REGION Network 141
   RUNG wire#powerrail
      Contact( "Carrier_06_Status.9" )
      Coil( "EMS".Carrier[06].SDC_IN.EncoderCommFault )
   END_RUNG
   // the same network as SCL:
   "EMS".Carrier[06].SDC_IN.EncoderCommFault := "Carrier_06_Status.9";
END_REGION

REGION Network 142
   RUNG wire#powerrail
      Contact( "Carrier_06_Status.10" )
      Coil( "EMS".Carrier[06].SDC_IN.DriveCommFault )
   END_RUNG
   // the same network as SCL:
   "EMS".Carrier[06].SDC_IN.DriveCommFault := "Carrier_06_Status.10";
END_REGION

REGION Network 143
   RUNG wire#powerrail
      Contact( "Carrier_06_Status.11" )
      Coil( "EMS".Carrier[06].SDC_IN.HMICommFault )
   END_RUNG
   // the same network as SCL:
   "EMS".Carrier[06].SDC_IN.HMICommFault := "Carrier_06_Status.11";
END_REGION

REGION Network 144
   RUNG wire#powerrail
      Contact( "Carrier_06_Status.2" )
      Coil( "EMS".Carrier[06].SDC_IN.AutoMode )
   END_RUNG
   RUNG wire#powerrail
      Contact( "Carrier_06_Status.1" )
      Coil( "EMS".Carrier[06].SDC_IN.ManualMode )
   END_RUNG
   // the same network as SCL:
   "EMS".Carrier[06].SDC_IN.AutoMode := "Carrier_06_Status.2";
   "EMS".Carrier[06].SDC_IN.ManualMode := "Carrier_06_Status.1";
END_REGION

REGION Network 145
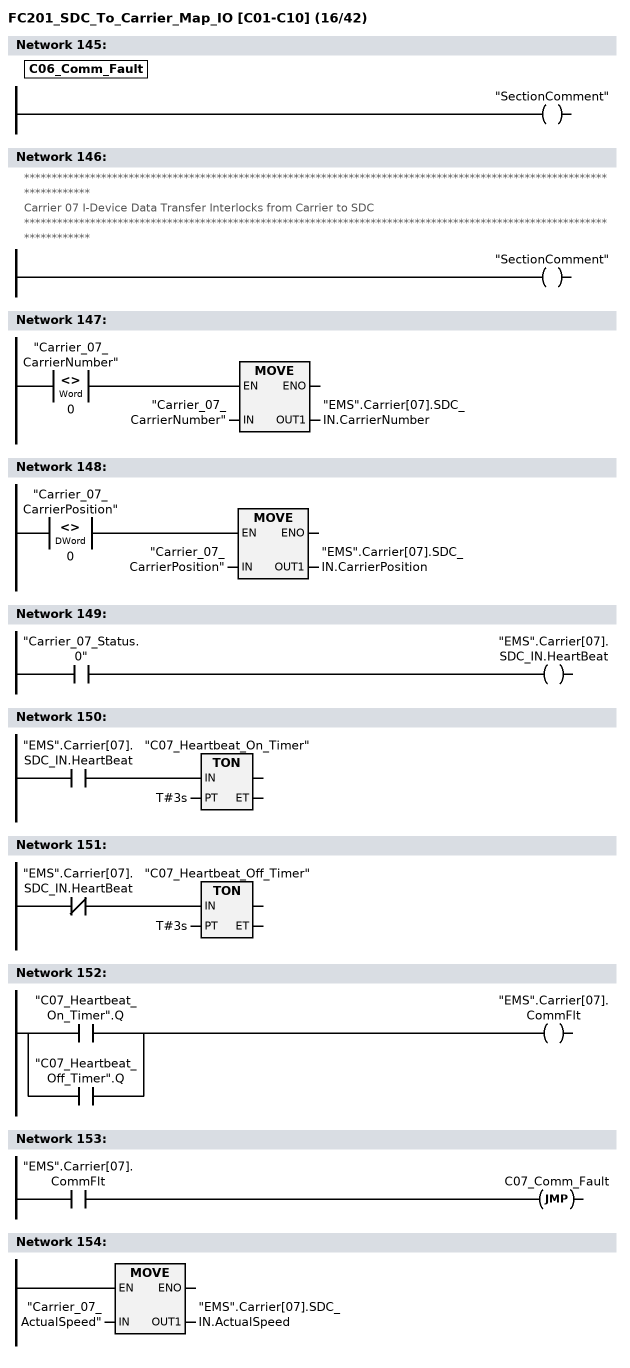
   Label( C06_Comm_Fault )
   RUNG wire#powerrail
      Coil( "SectionComment" )
   END_RUNG
   // the same network as SCL:
   C06_Comm_Fault:
   "SectionComment" := TRUE;
END_REGION

REGION Network 146
   // **********************************************************************************************************************
   // 
   // Carrier 07 I-Device Data Transfer Interlocks from Carrier to SDC
   // 
   // **********************************************************************************************************************
   RUNG wire#powerrail
      Coil( "SectionComment" )
   END_RUNG
   // the same network as SCL:
   "SectionComment" := TRUE;
END_REGION

REGION Network 147
   RUNG wire#powerrail
      { S7_Templates := "SrcType := Word" } NE_Contact(in1 := "Carrier_07_CarrierNumber", in2 := 0)
      Move(in := "Carrier_07_CarrierNumber", out1 => "EMS".Carrier[07].SDC_IN.CarrierNumber)
   END_RUNG
   // the same network as SCL:
   IF "Carrier_07_CarrierNumber" <> 0 THEN
       "EMS".Carrier[07].SDC_IN.CarrierNumber := "Carrier_07_CarrierNumber";
   END_IF;
END_REGION

REGION Network 148
   RUNG wire#powerrail
      { S7_Templates := "SrcType := DWord" } NE_Contact(in1 := "Carrier_07_CarrierPosition", in2 := 0)
      Move(in := "Carrier_07_CarrierPosition", out1 => "EMS".Carrier[07].SDC_IN.CarrierPosition)
   END_RUNG
   // the same network as SCL:
   IF "Carrier_07_CarrierPosition" <> 0 THEN
       "EMS".Carrier[07].SDC_IN.CarrierPosition := "Carrier_07_CarrierPosition";
   END_IF;
END_REGION

REGION Network 149
   RUNG wire#powerrail
      Contact( "Carrier_07_Status.0" )
      Coil( "EMS".Carrier[07].SDC_IN.HeartBeat )
   END_RUNG
   // the same network as SCL:
   "EMS".Carrier[07].SDC_IN.HeartBeat := "Carrier_07_Status.0";
END_REGION

REGION Network 150
   "C07_Heartbeat_On_Timer".TON(IN := "EMS".Carrier[07].SDC_IN.HeartBeat, PT := T#3s);
END_REGION

REGION Network 151
   "C07_Heartbeat_Off_Timer".TON(IN := NOT "EMS".Carrier[07].SDC_IN.HeartBeat, PT := T#3s);
END_REGION

REGION Network 152
   RUNG wire#powerrail
      Contact( "C07_Heartbeat_On_Timer".Q )
      wire#w1
      Coil( "EMS".Carrier[07].CommFlt )
   END_RUNG
   RUNG wire#powerrail
      Contact( "C07_Heartbeat_Off_Timer".Q )
   END_RUNG wire#w1
   // the same network as SCL:
   "EMS".Carrier[07].CommFlt := "C07_Heartbeat_On_Timer".Q OR "C07_Heartbeat_Off_Timer".Q;
END_REGION

REGION Network 153
   RUNG wire#powerrail
      Contact( "EMS".Carrier[07].CommFlt )
      JumpCoil( C07_Comm_Fault )
   END_RUNG
   // the same network as SCL:
   IF "EMS".Carrier[07].CommFlt THEN GOTO C07_Comm_Fault; END_IF;
END_REGION

REGION Network 154
   RUNG wire#powerrail
      Move(in := "Carrier_07_ActualSpeed", out1 => "EMS".Carrier[07].SDC_IN.ActualSpeed)
   END_RUNG
   // the same network as SCL:
   "EMS".Carrier[07].SDC_IN.ActualSpeed := "Carrier_07_ActualSpeed";
END_REGION

REGION Network 155
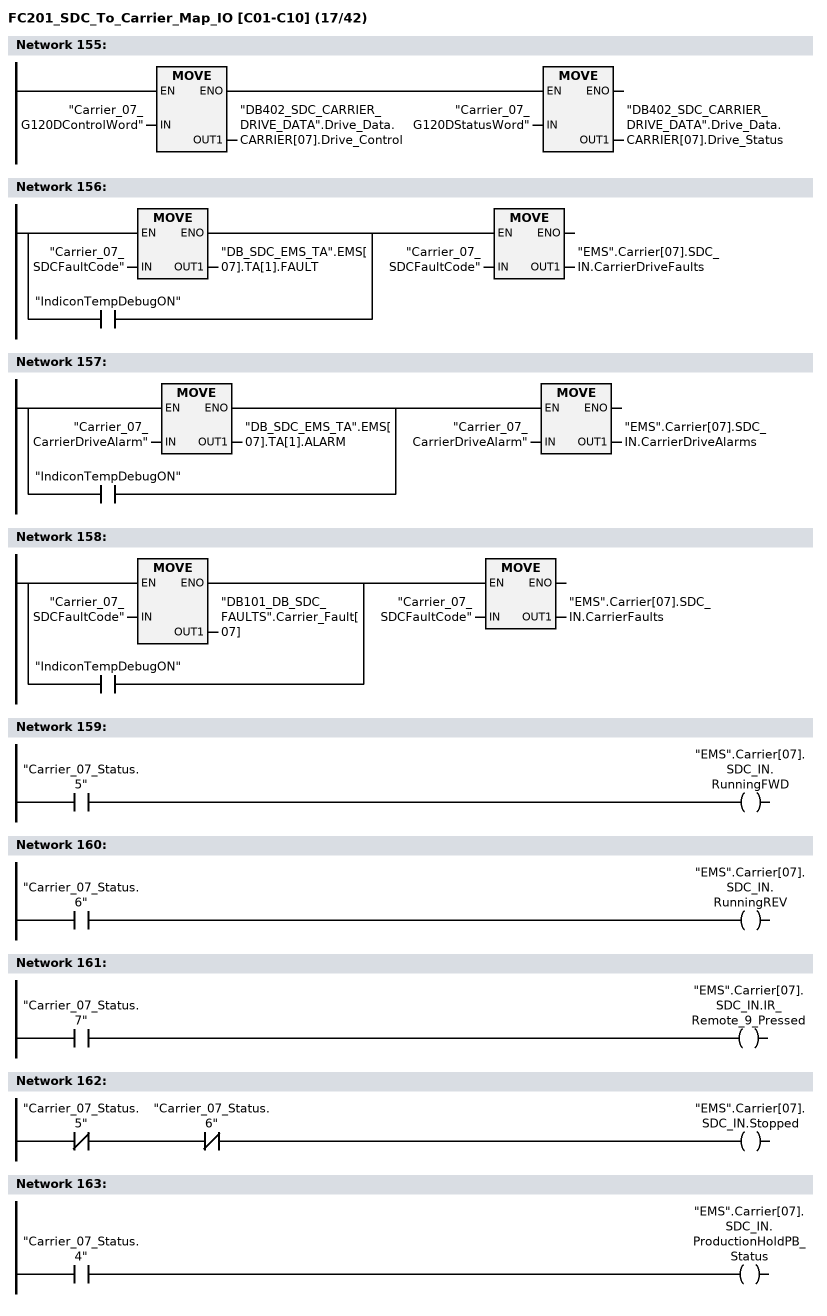
   RUNG wire#powerrail
      Move(in := "Carrier_07_G120DControlWord", out1 => "DB402_SDC_CARRIER_DRIVE_DATA".Drive_Data.CARRIER[07].Drive_Control)
      Move(in := "Carrier_07_G120DStatusWord", out1 => "DB402_SDC_CARRIER_DRIVE_DATA".Drive_Data.CARRIER[07].Drive_Status)
   END_RUNG
   // the same network as SCL:
   "DB402_SDC_CARRIER_DRIVE_DATA".Drive_Data.CARRIER[07].Drive_Control := "Carrier_07_G120DControlWord";
   "DB402_SDC_CARRIER_DRIVE_DATA".Drive_Data.CARRIER[07].Drive_Status := "Carrier_07_G120DStatusWord";
END_REGION

REGION Network 156
   RUNG wire#powerrail
      Move(in := "Carrier_07_SDCFaultCode", out1 => "DB_SDC_EMS_TA".EMS[07].TA[1].FAULT)
      wire#w1
      Move(in := "Carrier_07_SDCFaultCode", out1 => "EMS".Carrier[07].SDC_IN.CarrierDriveFaults)
   END_RUNG
   RUNG wire#powerrail
      Contact( "IndiconTempDebugON" )
   END_RUNG wire#w1
   // the same network as SCL:
   "DB_SDC_EMS_TA".EMS[07].TA[1].FAULT := "Carrier_07_SDCFaultCode";
   IF TRUE OR "IndiconTempDebugON" THEN
       "EMS".Carrier[07].SDC_IN.CarrierDriveFaults := "Carrier_07_SDCFaultCode";
   END_IF;
END_REGION

REGION Network 157
   RUNG wire#powerrail
      Move(in := "Carrier_07_CarrierDriveAlarm", out1 => "DB_SDC_EMS_TA".EMS[07].TA[1].ALARM)
      wire#w1
      Move(in := "Carrier_07_CarrierDriveAlarm", out1 => "EMS".Carrier[07].SDC_IN.CarrierDriveAlarms)
   END_RUNG
   RUNG wire#powerrail
      Contact( "IndiconTempDebugON" )
   END_RUNG wire#w1
   // the same network as SCL:
   "DB_SDC_EMS_TA".EMS[07].TA[1].ALARM := "Carrier_07_CarrierDriveAlarm";
   IF TRUE OR "IndiconTempDebugON" THEN
       "EMS".Carrier[07].SDC_IN.CarrierDriveAlarms := "Carrier_07_CarrierDriveAlarm";
   END_IF;
END_REGION

REGION Network 158
   RUNG wire#powerrail
      Move(in := "Carrier_07_SDCFaultCode", out1 => "DB101_DB_SDC_FAULTS".Carrier_Fault[07])
      wire#w1
      Move(in := "Carrier_07_SDCFaultCode", out1 => "EMS".Carrier[07].SDC_IN.CarrierFaults)
   END_RUNG
   RUNG wire#powerrail
      Contact( "IndiconTempDebugON" )
   END_RUNG wire#w1
   // the same network as SCL:
   "DB101_DB_SDC_FAULTS".Carrier_Fault[07] := "Carrier_07_SDCFaultCode";
   IF TRUE OR "IndiconTempDebugON" THEN
       "EMS".Carrier[07].SDC_IN.CarrierFaults := "Carrier_07_SDCFaultCode";
   END_IF;
END_REGION

REGION Network 159
   RUNG wire#powerrail
      Contact( "Carrier_07_Status.5" )
      Coil( "EMS".Carrier[07].SDC_IN.RunningFWD )
   END_RUNG
   // the same network as SCL:
   "EMS".Carrier[07].SDC_IN.RunningFWD := "Carrier_07_Status.5";
END_REGION

REGION Network 160
   RUNG wire#powerrail
      Contact( "Carrier_07_Status.6" )
      Coil( "EMS".Carrier[07].SDC_IN.RunningREV )
   END_RUNG
   // the same network as SCL:
   "EMS".Carrier[07].SDC_IN.RunningREV := "Carrier_07_Status.6";
END_REGION

REGION Network 161
   RUNG wire#powerrail
      Contact( "Carrier_07_Status.7" )
      Coil( "EMS".Carrier[07].SDC_IN.IR_Remote_9_Pressed )
   END_RUNG
   // the same network as SCL:
   "EMS".Carrier[07].SDC_IN.IR_Remote_9_Pressed := "Carrier_07_Status.7";
END_REGION

REGION Network 162
   RUNG wire#powerrail
      I_Contact( "Carrier_07_Status.5" )
      I_Contact( "Carrier_07_Status.6" )
      Coil( "EMS".Carrier[07].SDC_IN.Stopped )
   END_RUNG
   // the same network as SCL:
   "EMS".Carrier[07].SDC_IN.Stopped := NOT "Carrier_07_Status.5" AND NOT "Carrier_07_Status.6";
END_REGION

REGION Network 163
   RUNG wire#powerrail
      Contact( "Carrier_07_Status.4" )
      Coil( "EMS".Carrier[07].SDC_IN.ProductionHoldPB_Status )
   END_RUNG
   // the same network as SCL:
   "EMS".Carrier[07].SDC_IN.ProductionHoldPB_Status := "Carrier_07_Status.4";
END_REGION

REGION Network 164
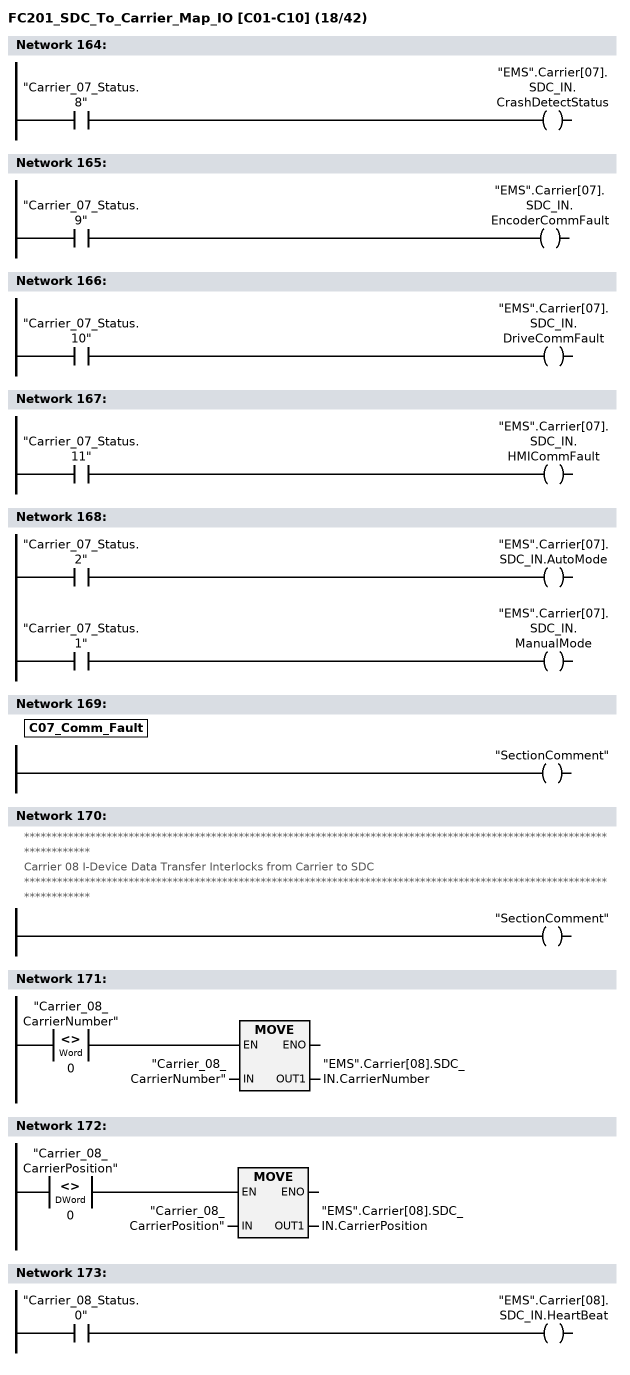
   RUNG wire#powerrail
      Contact( "Carrier_07_Status.8" )
      Coil( "EMS".Carrier[07].SDC_IN.CrashDetectStatus )
   END_RUNG
   // the same network as SCL:
   "EMS".Carrier[07].SDC_IN.CrashDetectStatus := "Carrier_07_Status.8";
END_REGION

REGION Network 165
   RUNG wire#powerrail
      Contact( "Carrier_07_Status.9" )
      Coil( "EMS".Carrier[07].SDC_IN.EncoderCommFault )
   END_RUNG
   // the same network as SCL:
   "EMS".Carrier[07].SDC_IN.EncoderCommFault := "Carrier_07_Status.9";
END_REGION

REGION Network 166
   RUNG wire#powerrail
      Contact( "Carrier_07_Status.10" )
      Coil( "EMS".Carrier[07].SDC_IN.DriveCommFault )
   END_RUNG
   // the same network as SCL:
   "EMS".Carrier[07].SDC_IN.DriveCommFault := "Carrier_07_Status.10";
END_REGION

REGION Network 167
   RUNG wire#powerrail
      Contact( "Carrier_07_Status.11" )
      Coil( "EMS".Carrier[07].SDC_IN.HMICommFault )
   END_RUNG
   // the same network as SCL:
   "EMS".Carrier[07].SDC_IN.HMICommFault := "Carrier_07_Status.11";
END_REGION

REGION Network 168
   RUNG wire#powerrail
      Contact( "Carrier_07_Status.2" )
      Coil( "EMS".Carrier[07].SDC_IN.AutoMode )
   END_RUNG
   RUNG wire#powerrail
      Contact( "Carrier_07_Status.1" )
      Coil( "EMS".Carrier[07].SDC_IN.ManualMode )
   END_RUNG
   // the same network as SCL:
   "EMS".Carrier[07].SDC_IN.AutoMode := "Carrier_07_Status.2";
   "EMS".Carrier[07].SDC_IN.ManualMode := "Carrier_07_Status.1";
END_REGION

REGION Network 169
   Label( C07_Comm_Fault )
   RUNG wire#powerrail
      Coil( "SectionComment" )
   END_RUNG
   // the same network as SCL:
   C07_Comm_Fault:
   "SectionComment" := TRUE;
END_REGION

REGION Network 170
   // **********************************************************************************************************************
   // 
   // Carrier 08 I-Device Data Transfer Interlocks from Carrier to SDC
   // 
   // **********************************************************************************************************************
   RUNG wire#powerrail
      Coil( "SectionComment" )
   END_RUNG
   // the same network as SCL:
   "SectionComment" := TRUE;
END_REGION

REGION Network 171
   RUNG wire#powerrail
      { S7_Templates := "SrcType := Word" } NE_Contact(in1 := "Carrier_08_CarrierNumber", in2 := 0)
      Move(in := "Carrier_08_CarrierNumber", out1 => "EMS".Carrier[08].SDC_IN.CarrierNumber)
   END_RUNG
   // the same network as SCL:
   IF "Carrier_08_CarrierNumber" <> 0 THEN
       "EMS".Carrier[08].SDC_IN.CarrierNumber := "Carrier_08_CarrierNumber";
   END_IF;
END_REGION

REGION Network 172
   RUNG wire#powerrail
      { S7_Templates := "SrcType := DWord" } NE_Contact(in1 := "Carrier_08_CarrierPosition", in2 := 0)
      Move(in := "Carrier_08_CarrierPosition", out1 => "EMS".Carrier[08].SDC_IN.CarrierPosition)
   END_RUNG
   // the same network as SCL:
   IF "Carrier_08_CarrierPosition" <> 0 THEN
       "EMS".Carrier[08].SDC_IN.CarrierPosition := "Carrier_08_CarrierPosition";
   END_IF;
END_REGION

REGION Network 173
   RUNG wire#powerrail
      Contact( "Carrier_08_Status.0" )
      Coil( "EMS".Carrier[08].SDC_IN.HeartBeat )
   END_RUNG
   // the same network as SCL:
   "EMS".Carrier[08].SDC_IN.HeartBeat := "Carrier_08_Status.0";
END_REGION

REGION Network 174
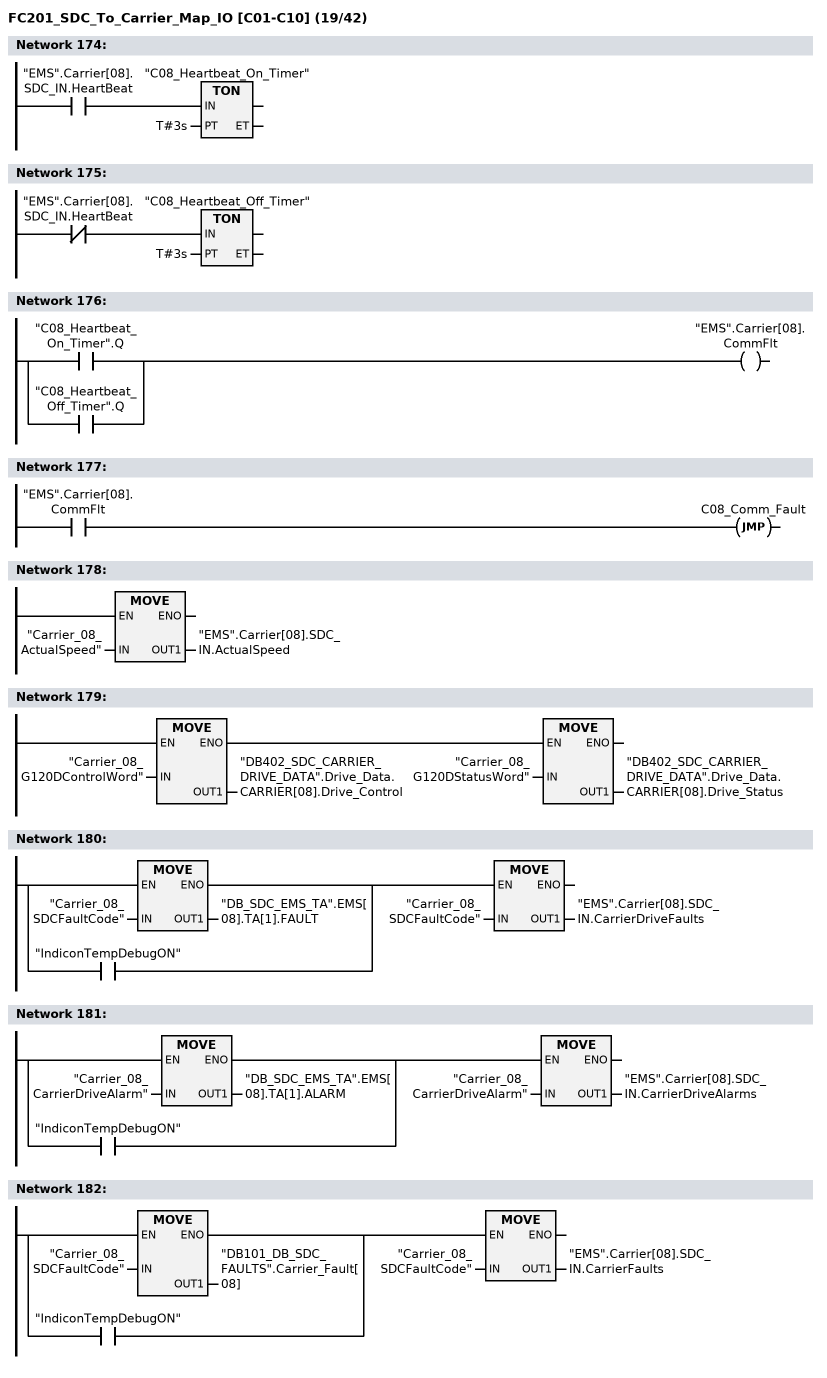
   "C08_Heartbeat_On_Timer".TON(IN := "EMS".Carrier[08].SDC_IN.HeartBeat, PT := T#3s);
END_REGION

REGION Network 175
   "C08_Heartbeat_Off_Timer".TON(IN := NOT "EMS".Carrier[08].SDC_IN.HeartBeat, PT := T#3s);
END_REGION

REGION Network 176
   RUNG wire#powerrail
      Contact( "C08_Heartbeat_On_Timer".Q )
      wire#w1
      Coil( "EMS".Carrier[08].CommFlt )
   END_RUNG
   RUNG wire#powerrail
      Contact( "C08_Heartbeat_Off_Timer".Q )
   END_RUNG wire#w1
   // the same network as SCL:
   "EMS".Carrier[08].CommFlt := "C08_Heartbeat_On_Timer".Q OR "C08_Heartbeat_Off_Timer".Q;
END_REGION

REGION Network 177
   RUNG wire#powerrail
      Contact( "EMS".Carrier[08].CommFlt )
      JumpCoil( C08_Comm_Fault )
   END_RUNG
   // the same network as SCL:
   IF "EMS".Carrier[08].CommFlt THEN GOTO C08_Comm_Fault; END_IF;
END_REGION

REGION Network 178
   RUNG wire#powerrail
      Move(in := "Carrier_08_ActualSpeed", out1 => "EMS".Carrier[08].SDC_IN.ActualSpeed)
   END_RUNG
   // the same network as SCL:
   "EMS".Carrier[08].SDC_IN.ActualSpeed := "Carrier_08_ActualSpeed";
END_REGION

REGION Network 179
   RUNG wire#powerrail
      Move(in := "Carrier_08_G120DControlWord", out1 => "DB402_SDC_CARRIER_DRIVE_DATA".Drive_Data.CARRIER[08].Drive_Control)
      Move(in := "Carrier_08_G120DStatusWord", out1 => "DB402_SDC_CARRIER_DRIVE_DATA".Drive_Data.CARRIER[08].Drive_Status)
   END_RUNG
   // the same network as SCL:
   "DB402_SDC_CARRIER_DRIVE_DATA".Drive_Data.CARRIER[08].Drive_Control := "Carrier_08_G120DControlWord";
   "DB402_SDC_CARRIER_DRIVE_DATA".Drive_Data.CARRIER[08].Drive_Status := "Carrier_08_G120DStatusWord";
END_REGION

REGION Network 180
   RUNG wire#powerrail
      Move(in := "Carrier_08_SDCFaultCode", out1 => "DB_SDC_EMS_TA".EMS[08].TA[1].FAULT)
      wire#w1
      Move(in := "Carrier_08_SDCFaultCode", out1 => "EMS".Carrier[08].SDC_IN.CarrierDriveFaults)
   END_RUNG
   RUNG wire#powerrail
      Contact( "IndiconTempDebugON" )
   END_RUNG wire#w1
   // the same network as SCL:
   "DB_SDC_EMS_TA".EMS[08].TA[1].FAULT := "Carrier_08_SDCFaultCode";
   IF TRUE OR "IndiconTempDebugON" THEN
       "EMS".Carrier[08].SDC_IN.CarrierDriveFaults := "Carrier_08_SDCFaultCode";
   END_IF;
END_REGION

REGION Network 181
   RUNG wire#powerrail
      Move(in := "Carrier_08_CarrierDriveAlarm", out1 => "DB_SDC_EMS_TA".EMS[08].TA[1].ALARM)
      wire#w1
      Move(in := "Carrier_08_CarrierDriveAlarm", out1 => "EMS".Carrier[08].SDC_IN.CarrierDriveAlarms)
   END_RUNG
   RUNG wire#powerrail
      Contact( "IndiconTempDebugON" )
   END_RUNG wire#w1
   // the same network as SCL:
   "DB_SDC_EMS_TA".EMS[08].TA[1].ALARM := "Carrier_08_CarrierDriveAlarm";
   IF TRUE OR "IndiconTempDebugON" THEN
       "EMS".Carrier[08].SDC_IN.CarrierDriveAlarms := "Carrier_08_CarrierDriveAlarm";
   END_IF;
END_REGION

REGION Network 182
   RUNG wire#powerrail
      Move(in := "Carrier_08_SDCFaultCode", out1 => "DB101_DB_SDC_FAULTS".Carrier_Fault[08])
      wire#w1
      Move(in := "Carrier_08_SDCFaultCode", out1 => "EMS".Carrier[08].SDC_IN.CarrierFaults)
   END_RUNG
   RUNG wire#powerrail
      Contact( "IndiconTempDebugON" )
   END_RUNG wire#w1
   // the same network as SCL:
   "DB101_DB_SDC_FAULTS".Carrier_Fault[08] := "Carrier_08_SDCFaultCode";
   IF TRUE OR "IndiconTempDebugON" THEN
       "EMS".Carrier[08].SDC_IN.CarrierFaults := "Carrier_08_SDCFaultCode";
   END_IF;
END_REGION

REGION Network 183
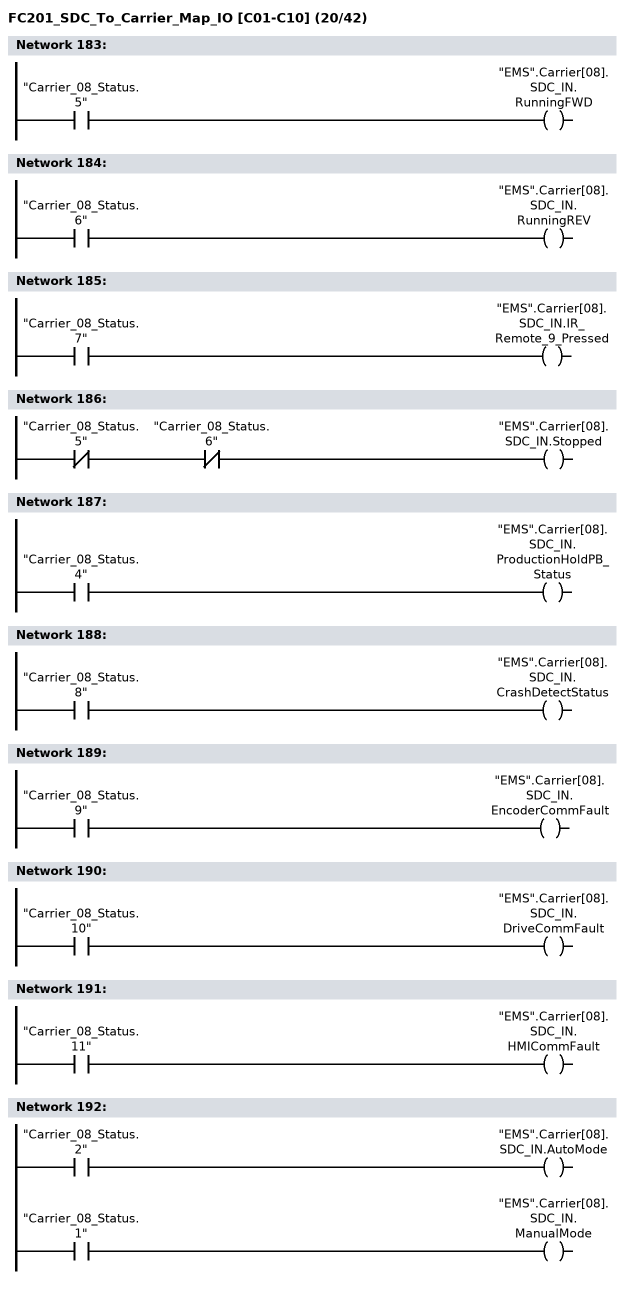
   RUNG wire#powerrail
      Contact( "Carrier_08_Status.5" )
      Coil( "EMS".Carrier[08].SDC_IN.RunningFWD )
   END_RUNG
   // the same network as SCL:
   "EMS".Carrier[08].SDC_IN.RunningFWD := "Carrier_08_Status.5";
END_REGION

REGION Network 184
   RUNG wire#powerrail
      Contact( "Carrier_08_Status.6" )
      Coil( "EMS".Carrier[08].SDC_IN.RunningREV )
   END_RUNG
   // the same network as SCL:
   "EMS".Carrier[08].SDC_IN.RunningREV := "Carrier_08_Status.6";
END_REGION

REGION Network 185
   RUNG wire#powerrail
      Contact( "Carrier_08_Status.7" )
      Coil( "EMS".Carrier[08].SDC_IN.IR_Remote_9_Pressed )
   END_RUNG
   // the same network as SCL:
   "EMS".Carrier[08].SDC_IN.IR_Remote_9_Pressed := "Carrier_08_Status.7";
END_REGION

REGION Network 186
   RUNG wire#powerrail
      I_Contact( "Carrier_08_Status.5" )
      I_Contact( "Carrier_08_Status.6" )
      Coil( "EMS".Carrier[08].SDC_IN.Stopped )
   END_RUNG
   // the same network as SCL:
   "EMS".Carrier[08].SDC_IN.Stopped := NOT "Carrier_08_Status.5" AND NOT "Carrier_08_Status.6";
END_REGION

REGION Network 187
   RUNG wire#powerrail
      Contact( "Carrier_08_Status.4" )
      Coil( "EMS".Carrier[08].SDC_IN.ProductionHoldPB_Status )
   END_RUNG
   // the same network as SCL:
   "EMS".Carrier[08].SDC_IN.ProductionHoldPB_Status := "Carrier_08_Status.4";
END_REGION

REGION Network 188
   RUNG wire#powerrail
      Contact( "Carrier_08_Status.8" )
      Coil( "EMS".Carrier[08].SDC_IN.CrashDetectStatus )
   END_RUNG
   // the same network as SCL:
   "EMS".Carrier[08].SDC_IN.CrashDetectStatus := "Carrier_08_Status.8";
END_REGION

REGION Network 189
   RUNG wire#powerrail
      Contact( "Carrier_08_Status.9" )
      Coil( "EMS".Carrier[08].SDC_IN.EncoderCommFault )
   END_RUNG
   // the same network as SCL:
   "EMS".Carrier[08].SDC_IN.EncoderCommFault := "Carrier_08_Status.9";
END_REGION

REGION Network 190
   RUNG wire#powerrail
      Contact( "Carrier_08_Status.10" )
      Coil( "EMS".Carrier[08].SDC_IN.DriveCommFault )
   END_RUNG
   // the same network as SCL:
   "EMS".Carrier[08].SDC_IN.DriveCommFault := "Carrier_08_Status.10";
END_REGION

REGION Network 191
   RUNG wire#powerrail
      Contact( "Carrier_08_Status.11" )
      Coil( "EMS".Carrier[08].SDC_IN.HMICommFault )
   END_RUNG
   // the same network as SCL:
   "EMS".Carrier[08].SDC_IN.HMICommFault := "Carrier_08_Status.11";
END_REGION

REGION Network 192
   RUNG wire#powerrail
      Contact( "Carrier_08_Status.2" )
      Coil( "EMS".Carrier[08].SDC_IN.AutoMode )
   END_RUNG
   RUNG wire#powerrail
      Contact( "Carrier_08_Status.1" )
      Coil( "EMS".Carrier[08].SDC_IN.ManualMode )
   END_RUNG
   // the same network as SCL:
   "EMS".Carrier[08].SDC_IN.AutoMode := "Carrier_08_Status.2";
   "EMS".Carrier[08].SDC_IN.ManualMode := "Carrier_08_Status.1";
END_REGION

REGION Network 193
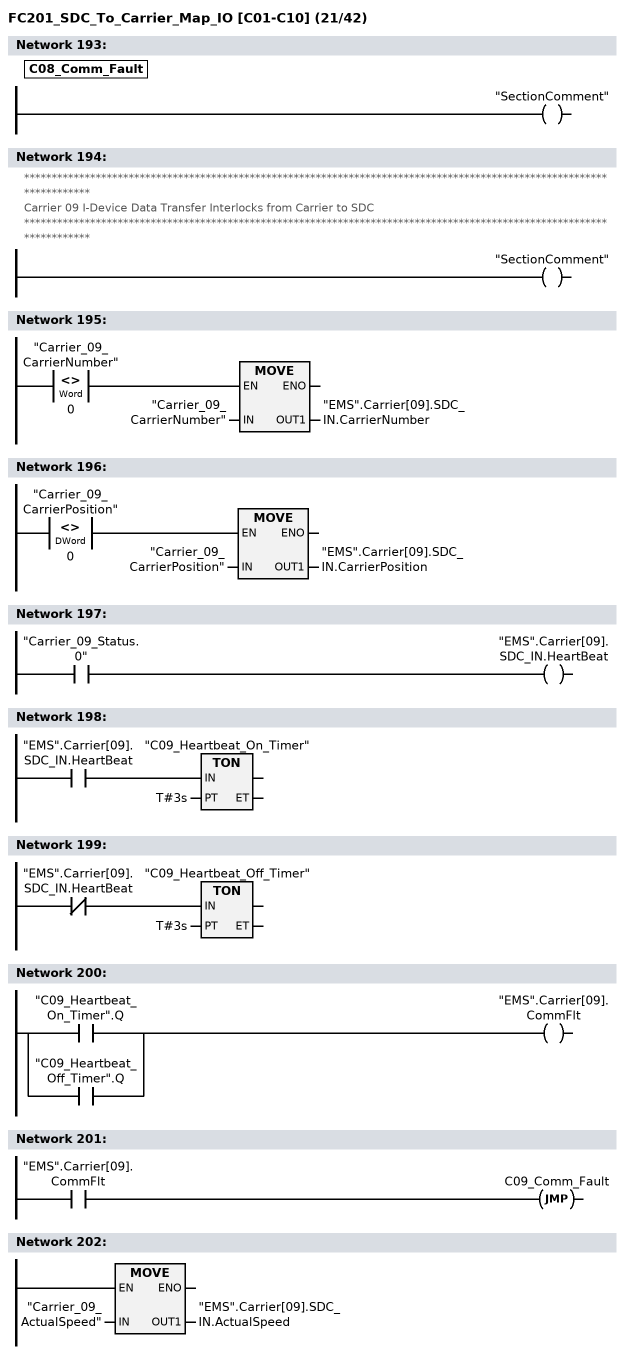
   Label( C08_Comm_Fault )
   RUNG wire#powerrail
      Coil( "SectionComment" )
   END_RUNG
   // the same network as SCL:
   C08_Comm_Fault:
   "SectionComment" := TRUE;
END_REGION

REGION Network 194
   // **********************************************************************************************************************
   // 
   // Carrier 09 I-Device Data Transfer Interlocks from Carrier to SDC
   // 
   // **********************************************************************************************************************
   RUNG wire#powerrail
      Coil( "SectionComment" )
   END_RUNG
   // the same network as SCL:
   "SectionComment" := TRUE;
END_REGION

REGION Network 195
   RUNG wire#powerrail
      { S7_Templates := "SrcType := Word" } NE_Contact(in1 := "Carrier_09_CarrierNumber", in2 := 0)
      Move(in := "Carrier_09_CarrierNumber", out1 => "EMS".Carrier[09].SDC_IN.CarrierNumber)
   END_RUNG
   // the same network as SCL:
   IF "Carrier_09_CarrierNumber" <> 0 THEN
       "EMS".Carrier[09].SDC_IN.CarrierNumber := "Carrier_09_CarrierNumber";
   END_IF;
END_REGION

REGION Network 196
   RUNG wire#powerrail
      { S7_Templates := "SrcType := DWord" } NE_Contact(in1 := "Carrier_09_CarrierPosition", in2 := 0)
      Move(in := "Carrier_09_CarrierPosition", out1 => "EMS".Carrier[09].SDC_IN.CarrierPosition)
   END_RUNG
   // the same network as SCL:
   IF "Carrier_09_CarrierPosition" <> 0 THEN
       "EMS".Carrier[09].SDC_IN.CarrierPosition := "Carrier_09_CarrierPosition";
   END_IF;
END_REGION

REGION Network 197
   RUNG wire#powerrail
      Contact( "Carrier_09_Status.0" )
      Coil( "EMS".Carrier[09].SDC_IN.HeartBeat )
   END_RUNG
   // the same network as SCL:
   "EMS".Carrier[09].SDC_IN.HeartBeat := "Carrier_09_Status.0";
END_REGION

REGION Network 198
   "C09_Heartbeat_On_Timer".TON(IN := "EMS".Carrier[09].SDC_IN.HeartBeat, PT := T#3s);
END_REGION

REGION Network 199
   "C09_Heartbeat_Off_Timer".TON(IN := NOT "EMS".Carrier[09].SDC_IN.HeartBeat, PT := T#3s);
END_REGION

REGION Network 200
   RUNG wire#powerrail
      Contact( "C09_Heartbeat_On_Timer".Q )
      wire#w1
      Coil( "EMS".Carrier[09].CommFlt )
   END_RUNG
   RUNG wire#powerrail
      Contact( "C09_Heartbeat_Off_Timer".Q )
   END_RUNG wire#w1
   // the same network as SCL:
   "EMS".Carrier[09].CommFlt := "C09_Heartbeat_On_Timer".Q OR "C09_Heartbeat_Off_Timer".Q;
END_REGION

REGION Network 201
   RUNG wire#powerrail
      Contact( "EMS".Carrier[09].CommFlt )
      JumpCoil( C09_Comm_Fault )
   END_RUNG
   // the same network as SCL:
   IF "EMS".Carrier[09].CommFlt THEN GOTO C09_Comm_Fault; END_IF;
END_REGION

REGION Network 202
   RUNG wire#powerrail
      Move(in := "Carrier_09_ActualSpeed", out1 => "EMS".Carrier[09].SDC_IN.ActualSpeed)
   END_RUNG
   // the same network as SCL:
   "EMS".Carrier[09].SDC_IN.ActualSpeed := "Carrier_09_ActualSpeed";
END_REGION

REGION Network 203
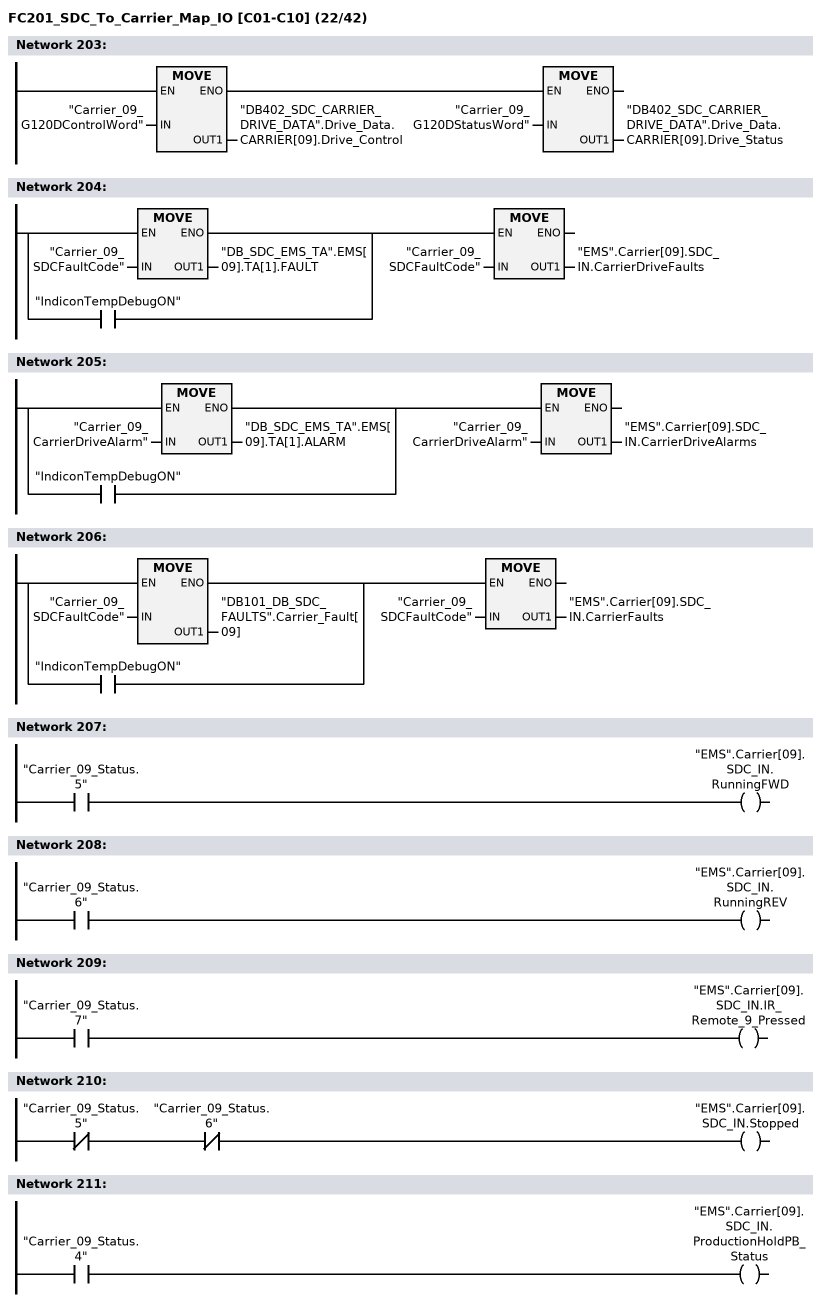
   RUNG wire#powerrail
      Move(in := "Carrier_09_G120DControlWord", out1 => "DB402_SDC_CARRIER_DRIVE_DATA".Drive_Data.CARRIER[09].Drive_Control)
      Move(in := "Carrier_09_G120DStatusWord", out1 => "DB402_SDC_CARRIER_DRIVE_DATA".Drive_Data.CARRIER[09].Drive_Status)
   END_RUNG
   // the same network as SCL:
   "DB402_SDC_CARRIER_DRIVE_DATA".Drive_Data.CARRIER[09].Drive_Control := "Carrier_09_G120DControlWord";
   "DB402_SDC_CARRIER_DRIVE_DATA".Drive_Data.CARRIER[09].Drive_Status := "Carrier_09_G120DStatusWord";
END_REGION

REGION Network 204
   RUNG wire#powerrail
      Move(in := "Carrier_09_SDCFaultCode", out1 => "DB_SDC_EMS_TA".EMS[09].TA[1].FAULT)
      wire#w1
      Move(in := "Carrier_09_SDCFaultCode", out1 => "EMS".Carrier[09].SDC_IN.CarrierDriveFaults)
   END_RUNG
   RUNG wire#powerrail
      Contact( "IndiconTempDebugON" )
   END_RUNG wire#w1
   // the same network as SCL:
   "DB_SDC_EMS_TA".EMS[09].TA[1].FAULT := "Carrier_09_SDCFaultCode";
   IF TRUE OR "IndiconTempDebugON" THEN
       "EMS".Carrier[09].SDC_IN.CarrierDriveFaults := "Carrier_09_SDCFaultCode";
   END_IF;
END_REGION

REGION Network 205
   RUNG wire#powerrail
      Move(in := "Carrier_09_CarrierDriveAlarm", out1 => "DB_SDC_EMS_TA".EMS[09].TA[1].ALARM)
      wire#w1
      Move(in := "Carrier_09_CarrierDriveAlarm", out1 => "EMS".Carrier[09].SDC_IN.CarrierDriveAlarms)
   END_RUNG
   RUNG wire#powerrail
      Contact( "IndiconTempDebugON" )
   END_RUNG wire#w1
   // the same network as SCL:
   "DB_SDC_EMS_TA".EMS[09].TA[1].ALARM := "Carrier_09_CarrierDriveAlarm";
   IF TRUE OR "IndiconTempDebugON" THEN
       "EMS".Carrier[09].SDC_IN.CarrierDriveAlarms := "Carrier_09_CarrierDriveAlarm";
   END_IF;
END_REGION

REGION Network 206
   RUNG wire#powerrail
      Move(in := "Carrier_09_SDCFaultCode", out1 => "DB101_DB_SDC_FAULTS".Carrier_Fault[09])
      wire#w1
      Move(in := "Carrier_09_SDCFaultCode", out1 => "EMS".Carrier[09].SDC_IN.CarrierFaults)
   END_RUNG
   RUNG wire#powerrail
      Contact( "IndiconTempDebugON" )
   END_RUNG wire#w1
   // the same network as SCL:
   "DB101_DB_SDC_FAULTS".Carrier_Fault[09] := "Carrier_09_SDCFaultCode";
   IF TRUE OR "IndiconTempDebugON" THEN
       "EMS".Carrier[09].SDC_IN.CarrierFaults := "Carrier_09_SDCFaultCode";
   END_IF;
END_REGION

REGION Network 207
   RUNG wire#powerrail
      Contact( "Carrier_09_Status.5" )
      Coil( "EMS".Carrier[09].SDC_IN.RunningFWD )
   END_RUNG
   // the same network as SCL:
   "EMS".Carrier[09].SDC_IN.RunningFWD := "Carrier_09_Status.5";
END_REGION

REGION Network 208
   RUNG wire#powerrail
      Contact( "Carrier_09_Status.6" )
      Coil( "EMS".Carrier[09].SDC_IN.RunningREV )
   END_RUNG
   // the same network as SCL:
   "EMS".Carrier[09].SDC_IN.RunningREV := "Carrier_09_Status.6";
END_REGION

REGION Network 209
   RUNG wire#powerrail
      Contact( "Carrier_09_Status.7" )
      Coil( "EMS".Carrier[09].SDC_IN.IR_Remote_9_Pressed )
   END_RUNG
   // the same network as SCL:
   "EMS".Carrier[09].SDC_IN.IR_Remote_9_Pressed := "Carrier_09_Status.7";
END_REGION

REGION Network 210
   RUNG wire#powerrail
      I_Contact( "Carrier_09_Status.5" )
      I_Contact( "Carrier_09_Status.6" )
      Coil( "EMS".Carrier[09].SDC_IN.Stopped )
   END_RUNG
   // the same network as SCL:
   "EMS".Carrier[09].SDC_IN.Stopped := NOT "Carrier_09_Status.5" AND NOT "Carrier_09_Status.6";
END_REGION

REGION Network 211
   RUNG wire#powerrail
      Contact( "Carrier_09_Status.4" )
      Coil( "EMS".Carrier[09].SDC_IN.ProductionHoldPB_Status )
   END_RUNG
   // the same network as SCL:
   "EMS".Carrier[09].SDC_IN.ProductionHoldPB_Status := "Carrier_09_Status.4";
END_REGION

REGION Network 212
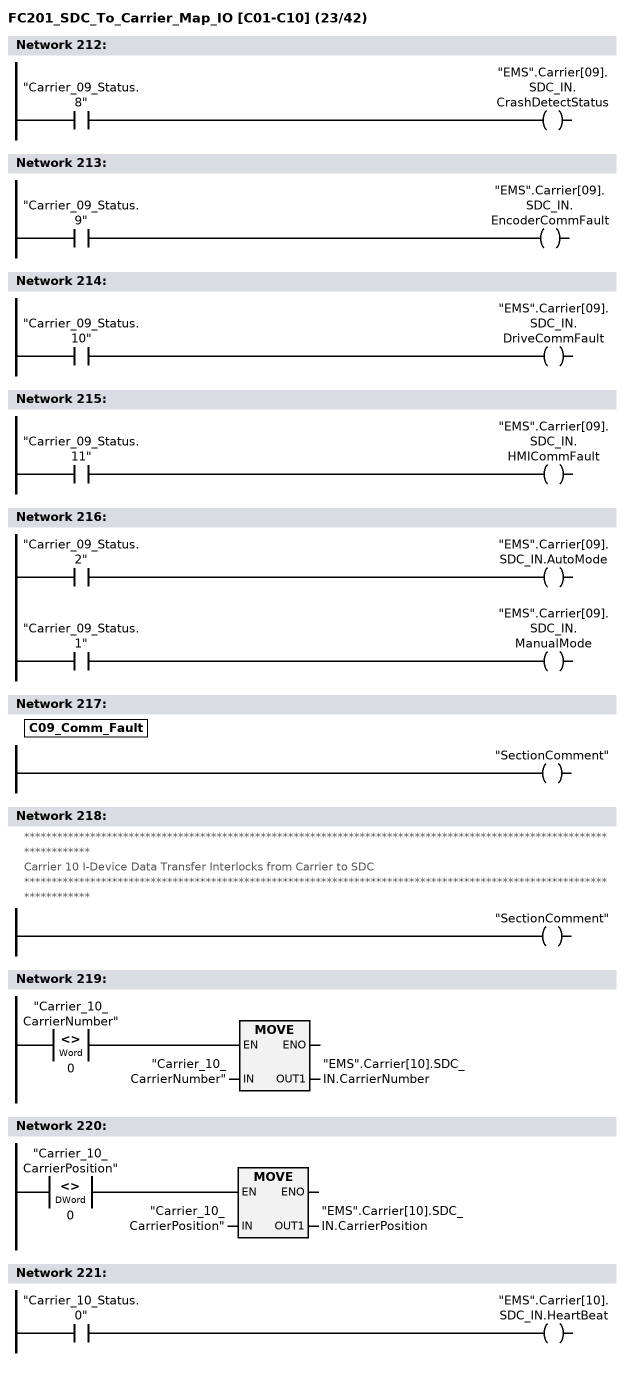
   RUNG wire#powerrail
      Contact( "Carrier_09_Status.8" )
      Coil( "EMS".Carrier[09].SDC_IN.CrashDetectStatus )
   END_RUNG
   // the same network as SCL:
   "EMS".Carrier[09].SDC_IN.CrashDetectStatus := "Carrier_09_Status.8";
END_REGION

REGION Network 213
   RUNG wire#powerrail
      Contact( "Carrier_09_Status.9" )
      Coil( "EMS".Carrier[09].SDC_IN.EncoderCommFault )
   END_RUNG
   // the same network as SCL:
   "EMS".Carrier[09].SDC_IN.EncoderCommFault := "Carrier_09_Status.9";
END_REGION

REGION Network 214
   RUNG wire#powerrail
      Contact( "Carrier_09_Status.10" )
      Coil( "EMS".Carrier[09].SDC_IN.DriveCommFault )
   END_RUNG
   // the same network as SCL:
   "EMS".Carrier[09].SDC_IN.DriveCommFault := "Carrier_09_Status.10";
END_REGION

REGION Network 215
   RUNG wire#powerrail
      Contact( "Carrier_09_Status.11" )
      Coil( "EMS".Carrier[09].SDC_IN.HMICommFault )
   END_RUNG
   // the same network as SCL:
   "EMS".Carrier[09].SDC_IN.HMICommFault := "Carrier_09_Status.11";
END_REGION

REGION Network 216
   RUNG wire#powerrail
      Contact( "Carrier_09_Status.2" )
      Coil( "EMS".Carrier[09].SDC_IN.AutoMode )
   END_RUNG
   RUNG wire#powerrail
      Contact( "Carrier_09_Status.1" )
      Coil( "EMS".Carrier[09].SDC_IN.ManualMode )
   END_RUNG
   // the same network as SCL:
   "EMS".Carrier[09].SDC_IN.AutoMode := "Carrier_09_Status.2";
   "EMS".Carrier[09].SDC_IN.ManualMode := "Carrier_09_Status.1";
END_REGION

REGION Network 217
   Label( C09_Comm_Fault )
   RUNG wire#powerrail
      Coil( "SectionComment" )
   END_RUNG
   // the same network as SCL:
   C09_Comm_Fault:
   "SectionComment" := TRUE;
END_REGION

REGION Network 218
   // **********************************************************************************************************************
   // 
   // Carrier 10 I-Device Data Transfer Interlocks from Carrier to SDC
   // 
   // **********************************************************************************************************************
   RUNG wire#powerrail
      Coil( "SectionComment" )
   END_RUNG
   // the same network as SCL:
   "SectionComment" := TRUE;
END_REGION

REGION Network 219
   RUNG wire#powerrail
      { S7_Templates := "SrcType := Word" } NE_Contact(in1 := "Carrier_10_CarrierNumber", in2 := 0)
      Move(in := "Carrier_10_CarrierNumber", out1 => "EMS".Carrier[10].SDC_IN.CarrierNumber)
   END_RUNG
   // the same network as SCL:
   IF "Carrier_10_CarrierNumber" <> 0 THEN
       "EMS".Carrier[10].SDC_IN.CarrierNumber := "Carrier_10_CarrierNumber";
   END_IF;
END_REGION

REGION Network 220
   RUNG wire#powerrail
      { S7_Templates := "SrcType := DWord" } NE_Contact(in1 := "Carrier_10_CarrierPosition", in2 := 0)
      Move(in := "Carrier_10_CarrierPosition", out1 => "EMS".Carrier[10].SDC_IN.CarrierPosition)
   END_RUNG
   // the same network as SCL:
   IF "Carrier_10_CarrierPosition" <> 0 THEN
       "EMS".Carrier[10].SDC_IN.CarrierPosition := "Carrier_10_CarrierPosition";
   END_IF;
END_REGION

REGION Network 221
   RUNG wire#powerrail
      Contact( "Carrier_10_Status.0" )
      Coil( "EMS".Carrier[10].SDC_IN.HeartBeat )
   END_RUNG
   // the same network as SCL:
   "EMS".Carrier[10].SDC_IN.HeartBeat := "Carrier_10_Status.0";
END_REGION

REGION Network 222
